   "EMP IDB_stations_me{16}_partNumbers{2}" : WString[40] = PLC "EMP IDB".stations.me[16].partNumbers[2], 1 s
   "EMP IDB_stations_me{16}_partNumbers{3}" : WString[40] = PLC "EMP IDB".stations.me[16].partNumbers[3], 1 s
   "EMP IDB_stations_me{16}_partNumbers{4}" : WString[40] = PLC "EMP IDB".stations.me[16].partNumbers[4], 1 s
   "EMP IDB_stations_me{16}_partNumbers{5}" : WString[40] = PLC "EMP IDB".stations.me[16].partNumbers[5], 1 s
   "EMP IDB_stations_me{16}_partNumbers{6}" : WString[40] = PLC "EMP IDB".stations.me[16].partNumbers[6], 1 s
   "EMP IDB_stations_me{16}_partNumbers{7}" : WString[40] = PLC "EMP IDB".stations.me[16].partNumbers[7], 1 s
   "EMP IDB_stations_me{17}_partNumbers{0}" : WString[40] = PLC "EMP IDB".stations.me[17].partNumbers[0], 1 s
   "EMP IDB_stations_me{17}_partNumbers{1}" : WString[40] = PLC "EMP IDB".stations.me[17].partNumbers[1], 1 s
   "EMP IDB_stations_me{17}_partNumbers{2}" : WString[40] = PLC "EMP IDB".stations.me[17].partNumbers[2], 1 s
   "EMP IDB_stations_me{17}_partNumbers{3}" : WString[40] = PLC "EMP IDB".stations.me[17].partNumbers[3], 1 s
   "EMP IDB_stations_me{17}_partNumbers{4}" : WString[40] = PLC "EMP IDB".stations.me[17].partNumbers[4], 1 s
   "EMP IDB_stations_me{17}_partNumbers{5}" : WString[40] = PLC "EMP IDB".stations.me[17].partNumbers[5], 1 s
   "EMP IDB_stations_me{17}_partNumbers{6}" : WString[40] = PLC "EMP IDB".stations.me[17].partNumbers[6], 1 s
   "EMP IDB_stations_me{17}_partNumbers{7}" : WString[40] = PLC "EMP IDB".stations.me[17].partNumbers[7], 1 s
   "EMP IDB_stations_me{18}_partNumbers{0}" : WString[40] = PLC "EMP IDB".stations.me[18].partNumbers[0], 1 s
   "EMP IDB_stations_me{18}_partNumbers{1}" : WString[40] = PLC "EMP IDB".stations.me[18].partNumbers[1], 1 s
   "EMP IDB_stations_me{18}_partNumbers{2}" : WString[40] = PLC "EMP IDB".stations.me[18].partNumbers[2], 1 s
   "EMP IDB_stations_me{18}_partNumbers{3}" : WString[40] = PLC "EMP IDB".stations.me[18].partNumbers[3], 1 s
   "EMP IDB_stations_me{18}_partNumbers{4}" : WString[40] = PLC "EMP IDB".stations.me[18].partNumbers[4], 1 s
   "EMP IDB_stations_me{18}_partNumbers{5}" : WString[40] = PLC "EMP IDB".stations.me[18].partNumbers[5], 1 s
   "EMP IDB_stations_me{18}_partNumbers{6}" : WString[40] = PLC "EMP IDB".stations.me[18].partNumbers[6], 1 s
   "EMP IDB_stations_me{18}_partNumbers{7}" : WString[40] = PLC "EMP IDB".stations.me[18].partNumbers[7], 1 s
   "EMP IDB_stations_me{19}_partNumbers{0}" : WString[40] = PLC "EMP IDB".stations.me[19].partNumbers[0], 1 s
   "EMP IDB_stations_me{19}_partNumbers{1}" : WString[40] = PLC "EMP IDB".stations.me[19].partNumbers[1], 1 s
   "EMP IDB_stations_me{19}_partNumbers{2}" : WString[40] = PLC "EMP IDB".stations.me[19].partNumbers[2], 1 s
   "EMP IDB_stations_me{19}_partNumbers{3}" : WString[40] = PLC "EMP IDB".stations.me[19].partNumbers[3], 1 s
   "EMP IDB_stations_me{19}_partNumbers{4}" : WString[40] = PLC "EMP IDB".stations.me[19].partNumbers[4], 1 s
   "EMP IDB_stations_me{19}_partNumbers{5}" : WString[40] = PLC "EMP IDB".stations.me[19].partNumbers[5], 1 s
   "EMP IDB_stations_me{19}_partNumbers{6}" : WString[40] = PLC "EMP IDB".stations.me[19].partNumbers[6], 1 s
   "EMP IDB_stations_me{19}_partNumbers{7}" : WString[40] = PLC "EMP IDB".stations.me[19].partNumbers[7], 1 s
   "EMP IDB_stations_me{20}_partNumbers{0}" : WString[40] = PLC "EMP IDB".stations.me[20].partNumbers[0], 1 s
   "EMP IDB_stations_me{20}_partNumbers{1}" : WString[40] = PLC "EMP IDB".stations.me[20].partNumbers[1], 1 s
   "EMP IDB_stations_me{20}_partNumbers{2}" : WString[40] = PLC "EMP IDB".stations.me[20].partNumbers[2], 1 s
   "EMP IDB_stations_me{20}_partNumbers{3}" : WString[40] = PLC "EMP IDB".stations.me[20].partNumbers[3], 1 s
   "EMP IDB_stations_me{20}_partNumbers{4}" : WString[40] = PLC "EMP IDB".stations.me[20].partNumbers[4], 1 s
   "EMP IDB_stations_me{20}_partNumbers{5}" : WString[40] = PLC "EMP IDB".stations.me[20].partNumbers[5], 1 s
   "EMP IDB_stations_me{20}_partNumbers{6}" : WString[40] = PLC "EMP IDB".stations.me[20].partNumbers[6], 1 s
   "EMP IDB_stations_me{20}_partNumbers{7}" : WString[40] = PLC "EMP IDB".stations.me[20].partNumbers[7], 1 s
   "EMP IDB_stations_me{21}_partNumbers{0}" : WString[40] = PLC "EMP IDB".stations.me[21].partNumbers[0], 1 s
   "EMP IDB_stations_me{21}_partNumbers{1}" : WString[40] = PLC "EMP IDB".stations.me[21].partNumbers[1], 1 s
   "EMP IDB_stations_me{21}_partNumbers{2}" : WString[40] = PLC "EMP IDB".stations.me[21].partNumbers[2], 1 s
   "EMP IDB_stations_me{21}_partNumbers{3}" : WString[40] = PLC "EMP IDB".stations.me[21].partNumbers[3], 1 s
   "EMP IDB_stations_me{21}_partNumbers{4}" : WString[40] = PLC "EMP IDB".stations.me[21].partNumbers[4], 1 s
   "EMP IDB_stations_me{21}_partNumbers{5}" : WString[40] = PLC "EMP IDB".stations.me[21].partNumbers[5], 1 s
   "EMP IDB_stations_me{21}_partNumbers{6}" : WString[40] = PLC "EMP IDB".stations.me[21].partNumbers[6], 1 s
   "EMP IDB_stations_me{21}_partNumbers{7}" : WString[40] = PLC "EMP IDB".stations.me[21].partNumbers[7], 1 s
   "EMP IDB_stations_me{22}_partNumbers{0}" : WString[40] = PLC "EMP IDB".stations.me[22].partNumbers[0], 1 s
   "EMP IDB_stations_me{22}_partNumbers{1}" : WString[40] = PLC "EMP IDB".stations.me[22].partNumbers[1], 1 s
   "EMP IDB_stations_me{22}_partNumbers{2}" : WString[40] = PLC "EMP IDB".stations.me[22].partNumbers[2], 1 s
   "EMP IDB_stations_me{22}_partNumbers{3}" : WString[40] = PLC "EMP IDB".stations.me[22].partNumbers[3], 1 s
   "EMP IDB_stations_me{22}_partNumbers{4}" : WString[40] = PLC "EMP IDB".stations.me[22].partNumbers[4], 1 s
   "EMP IDB_stations_me{22}_partNumbers{5}" : WString[40] = PLC "EMP IDB".stations.me[22].partNumbers[5], 1 s
   "EMP IDB_stations_me{22}_partNumbers{6}" : WString[40] = PLC "EMP IDB".stations.me[22].partNumbers[6], 1 s
   "EMP IDB_stations_me{22}_partNumbers{7}" : WString[40] = PLC "EMP IDB".stations.me[22].partNumbers[7], 1 s
   "EMP IDB_stations_me{23}_partNumbers{0}" : WString[40] = PLC "EMP IDB".stations.me[23].partNumbers[0], 1 s
   "EMP IDB_stations_me{23}_partNumbers{1}" : WString[40] = PLC "EMP IDB".stations.me[23].partNumbers[1], 1 s
   "EMP IDB_stations_me{23}_partNumbers{2}" : WString[40] = PLC "EMP IDB".stations.me[23].partNumbers[2], 1 s
   "EMP IDB_stations_me{23}_partNumbers{3}" : WString[40] = PLC "EMP IDB".stations.me[23].partNumbers[3], 1 s
   "EMP IDB_stations_me{23}_partNumbers{4}" : WString[40] = PLC "EMP IDB".stations.me[23].partNumbers[4], 1 s
   "EMP IDB_stations_me{23}_partNumbers{5}" : WString[40] = PLC "EMP IDB".stations.me[23].partNumbers[5], 1 s
   "EMP IDB_stations_me{23}_partNumbers{6}" : WString[40] = PLC "EMP IDB".stations.me[23].partNumbers[6], 1 s
   "EMP IDB_stations_me{23}_partNumbers{7}" : WString[40] = PLC "EMP IDB".stations.me[23].partNumbers[7], 1 s
   "EMP IDB_stations_me{3}_partNumbers{0}" : WString[40] = PLC "EMP IDB".stations.me[3].partNumbers[0], 1 s

text list "Station Selection Single": 0 'Select a Station to View'; 1 'Assignments'

recipe "VOLVO 16 01": Button 0 <- "EMP IDB_stations_me{0}_partNumbers{0}", Button 1 <- "EMP IDB_stations_me{0}_partNumbers{1}", Button 2 <- "EMP IDB_stations_me{0}_partNumbers{2}", Button 3 <- "EMP IDB_stations_me{0}_partNumbers{3}", Button 4 <- "EMP IDB_stations_me{0}_partNumbers{4}", Button 5 <- "EMP IDB_stations_me{0}_partNumbers{5}", Button 6 <- "EMP IDB_stations_me{0}_partNumbers{6}", Button 7 <- "EMP IDB_stations_me{0}_partNumbers{7}"

recipe "VOLVO 16 02": Button 0 <- "EMP IDB_stations_me{1}_partNumbers{0}", Button 1 <- "EMP IDB_stations_me{1}_partNumbers{1}", Button 2 <- "EMP IDB_stations_me{1}_partNumbers{2}", Button 3 <- "EMP IDB_stations_me{1}_partNumbers{3}", Button 4 <- "EMP IDB_stations_me{1}_partNumbers{4}", Button 5 <- "EMP IDB_stations_me{1}_partNumbers{5}", Button 6 <- "EMP IDB_stations_me{1}_partNumbers{6}", Button 7 <- "EMP IDB_stations_me{1}_partNumbers{7}"

recipe "VOLVO 16 03": Button 0 <- "EMP IDB_stations_me{2}_partNumbers{0}", Button 1 <- "EMP IDB_stations_me{2}_partNumbers{1}", Button 2 <- "EMP IDB_stations_me{2}_partNumbers{2}", Button 3 <- "EMP IDB_stations_me{2}_partNumbers{3}", Button 4 <- "EMP IDB_stations_me{2}_partNumbers{4}", Button 5 <- "EMP IDB_stations_me{2}_partNumbers{5}", Button 6 <- "EMP IDB_stations_me{2}_partNumbers{6}", Button 7 <- "EMP IDB_stations_me{2}_partNumbers{7}"

recipe "VOLVO 16 04": Button 0 <- "EMP IDB_stations_me{3}_partNumbers{0}", Button 1, Button 2, Button 3, Button 4, Button 5, Button 6, Button 7, Recipe_element_1

recipe "VOLVO 16 05": Button 0 <- "EMP IDB_stations_me{4}_partNumbers{0}", Button 1 <- "EMP IDB_stations_me{4}_partNumbers{1}", Button 2 <- "EMP IDB_stations_me{4}_partNumbers{2}", Button 3 <- "EMP IDB_stations_me{4}_partNumbers{3}", Button 4 <- "EMP IDB_stations_me{4}_partNumbers{4}", Button 5 <- "EMP IDB_stations_me{4}_partNumbers{5}", Button 6 <- "EMP IDB_stations_me{4}_partNumbers{6}", Button 7 <- "EMP IDB_stations_me{4}_partNumbers{7}"

recipe "VOLVO 16 06": Button 0 <- "EMP IDB_stations_me{5}_partNumbers{0}", Button 1 <- "EMP IDB_stations_me{5}_partNumbers{1}", Button 2 <- "EMP IDB_stations_me{5}_partNumbers{2}", Button 3 <- "EMP IDB_stations_me{5}_partNumbers{3}", Button 4 <- "EMP IDB_stations_me{5}_partNumbers{4}", Button 5 <- "EMP IDB_stations_me{5}_partNumbers{5}", Button 6 <- "EMP IDB_stations_me{5}_partNumbers{6}", Button 7 <- "EMP IDB_stations_me{5}_partNumbers{7}"

recipe "VOLVO 16 07": Button 0 <- "EMP IDB_stations_me{6}_partNumbers{0}", Button 1 <- "EMP IDB_stations_me{6}_partNumbers{1}", Button 2 <- "EMP IDB_stations_me{6}_partNumbers{2}", Button 3 <- "EMP IDB_stations_me{6}_partNumbers{3}", Button 4 <- "EMP IDB_stations_me{6}_partNumbers{4}", Button 5 <- "EMP IDB_stations_me{6}_partNumbers{5}", Button 6 <- "EMP IDB_stations_me{6}_partNumbers{6}", Button 7 <- "EMP IDB_stations_me{6}_partNumbers{7}"

recipe "VOLVO 16 08": Button 0 <- "EMP IDB_stations_me{7}_partNumbers{0}", Button 1 <- "EMP IDB_stations_me{7}_partNumbers{1}", Button 2 <- "EMP IDB_stations_me{7}_partNumbers{2}", Button 3 <- "EMP IDB_stations_me{7}_partNumbers{3}", Button 4 <- "EMP IDB_stations_me{7}_partNumbers{4}", Button 5 <- "EMP IDB_stations_me{7}_partNumbers{5}", Button 6 <- "EMP IDB_stations_me{7}_partNumbers{6}", Button 7 <- "EMP IDB_stations_me{7}_partNumbers{7}"

recipe "VOLVO 16 09": Button 0 <- "EMP IDB_stations_me{8}_partNumbers{0}", Button 1 <- "EMP IDB_stations_me{8}_partNumbers{1}", Button 2 <- "EMP IDB_stations_me{8}_partNumbers{2}", Button 3 <- "EMP IDB_stations_me{8}_partNumbers{3}", Button 4 <- "EMP IDB_stations_me{8}_partNumbers{4}", Button 5 <- "EMP IDB_stations_me{8}_partNumbers{5}", Button 6 <- "EMP IDB_stations_me{8}_partNumbers{6}", Button 7 <- "EMP IDB_stations_me{8}_partNumbers{7}"

recipe "VOLVO 16 10": Button 0 <- "EMP IDB_stations_me{9}_partNumbers{0}", Button 1 <- "EMP IDB_stations_me{9}_partNumbers{1}", Button 2 <- "EMP IDB_stations_me{9}_partNumbers{2}", Button 3 <- "EMP IDB_stations_me{9}_partNumbers{3}", Button 4 <- "EMP IDB_stations_me{9}_partNumbers{4}", Button 5 <- "EMP IDB_stations_me{9}_partNumbers{5}", Button 6 <- "EMP IDB_stations_me{9}_partNumbers{6}", Button 7 <- "EMP IDB_stations_me{9}_partNumbers{7}"

recipe "VOLVO 16 11": Button 0 <- "EMP IDB_stations_me{10}_partNumbers{0}", Button 1 <- "EMP IDB_stations_me{10}_partNumbers{1}", Button 2 <- "EMP IDB_stations_me{10}_partNumbers{2}", Button 3 <- "EMP IDB_stations_me{10}_partNumbers{3}", Button 4 <- "EMP IDB_stations_me{10}_partNumbers{4}", Button 5 <- "EMP IDB_stations_me{10}_partNumbers{5}", Button 6 <- "EMP IDB_stations_me{10}_partNumbers{6}", Button 7 <- "EMP IDB_stations_me{10}_partNumbers{7}"

recipe "CHM 01": Button 0 <- "EMP IDB_stations_me{11}_partNumbers{0}", Button 1 <- "EMP IDB_stations_me{11}_partNumbers{1}", Button 2 <- "EMP IDB_stations_me{11}_partNumbers{2}", Button 3 <- "EMP IDB_stations_me{11}_partNumbers{3}", Button 4 <- "EMP IDB_stations_me{11}_partNumbers{4}", Button 5 <- "EMP IDB_stations_me{11}_partNumbers{5}", Button 6 <- "EMP IDB_stations_me{11}_partNumbers{6}", Button 7 <- "EMP IDB_stations_me{11}_partNumbers{7}"

recipe "CHM 02": Button 0 <- "EMP IDB_stations_me{12}_partNumbers{0}", Button 1 <- "EMP IDB_stations_me{12}_partNumbers{1}", Button 2 <- "EMP IDB_stations_me{12}_partNumbers{2}", Button 3 <- "EMP IDB_stations_me{12}_partNumbers{3}", Button 4 <- "EMP IDB_stations_me{12}_partNumbers{4}", Button 5 <- "EMP IDB_stations_me{12}_partNumbers{5}", Button 6 <- "EMP IDB_stations_me{12}_partNumbers{6}", Button 7 <- "EMP IDB_stations_me{12}_partNumbers{7}"

recipe "CHM 03": Button 0 <- "EMP IDB_stations_me{13}_partNumbers{0}", Button 1 <- "EMP IDB_stations_me{13}_partNumbers{1}", Button 2 <- "EMP IDB_stations_me{13}_partNumbers{2}", Button 3 <- "EMP IDB_stations_me{13}_partNumbers{3}", Button 4 <- "EMP IDB_stations_me{13}_partNumbers{4}", Button 5 <- "EMP IDB_stations_me{13}_partNumbers{5}", Button 6 <- "EMP IDB_stations_me{13}_partNumbers{6}", Button 7 <- "EMP IDB_stations_me{13}_partNumbers{7}"

recipe "CHM 04": Button 0 <- "EMP IDB_stations_me{14}_partNumbers{0}", Button 1 <- "EMP IDB_stations_me{14}_partNumbers{1}", Button 2 <- "EMP IDB_stations_me{14}_partNumbers{2}", Button 3 <- "EMP IDB_stations_me{14}_partNumbers{3}", Button 4 <- "EMP IDB_stations_me{14}_partNumbers{4}", Button 5 <- "EMP IDB_stations_me{14}_partNumbers{5}", Button 6 <- "EMP IDB_stations_me{14}_partNumbers{6}", Button 7 <- "EMP IDB_stations_me{14}_partNumbers{7}"

recipe "CHM 05": Button 0 <- "EMP IDB_stations_me{15}_partNumbers{0}", Button 1 <- "EMP IDB_stations_me{15}_partNumbers{1}", Button 2 <- "EMP IDB_stations_me{15}_partNumbers{2}", Button 3 <- "EMP IDB_stations_me{15}_partNumbers{3}", Button 4 <- "EMP IDB_stations_me{15}_partNumbers{4}", Button 5 <- "EMP IDB_stations_me{15}_partNumbers{5}", Button 6 <- "EMP IDB_stations_me{15}_partNumbers{6}", Button 7 <- "EMP IDB_stations_me{15}_partNumbers{7}"

recipe "CDO 01": Button 0 <- "EMP IDB_stations_me{16}_partNumbers{0}", Button 1 <- "EMP IDB_stations_me{16}_partNumbers{1}", Button 2 <- "EMP IDB_stations_me{16}_partNumbers{2}", Button 3 <- "EMP IDB_stations_me{16}_partNumbers{3}", Button 4 <- "EMP IDB_stations_me{16}_partNumbers{4}", Button 5 <- "EMP IDB_stations_me{16}_partNumbers{5}", Button 6 <- "EMP IDB_stations_me{16}_partNumbers{6}", Button 7 <- "EMP IDB_stations_me{16}_partNumbers{7}"

recipe "CDO 02": Button 0 <- "EMP IDB_stations_me{17}_partNumbers{0}", Button 1 <- "EMP IDB_stations_me{17}_partNumbers{1}", Button 2 <- "EMP IDB_stations_me{17}_partNumbers{2}", Button 3 <- "EMP IDB_stations_me{17}_partNumbers{3}", Button 4 <- "EMP IDB_stations_me{17}_partNumbers{4}", Button 5 <- "EMP IDB_stations_me{17}_partNumbers{5}", Button 6 <- "EMP IDB_stations_me{17}_partNumbers{6}", Button 7 <- "EMP IDB_stations_me{17}_partNumbers{7}"

recipe "CDO 03": Button 0 <- "EMP IDB_stations_me{18}_partNumbers{0}", Button 1 <- "EMP IDB_stations_me{18}_partNumbers{1}", Button 2 <- "EMP IDB_stations_me{18}_partNumbers{2}", Button 3 <- "EMP IDB_stations_me{18}_partNumbers{3}", Button 4 <- "EMP IDB_stations_me{18}_partNumbers{4}", Button 5 <- "EMP IDB_stations_me{18}_partNumbers{5}", Button 6 <- "EMP IDB_stations_me{18}_partNumbers{6}", Button 7 <- "EMP IDB_stations_me{18}_partNumbers{7}"

recipe "BFL 01": Button 0 <- "EMP IDB_stations_me{19}_partNumbers{0}", Button 1 <- "EMP IDB_stations_me{19}_partNumbers{1}", Button 2 <- "EMP IDB_stations_me{19}_partNumbers{2}", Button 3 <- "EMP IDB_stations_me{19}_partNumbers{3}", Button 4 <- "EMP IDB_stations_me{19}_partNumbers{4}", Button 5 <- "EMP IDB_stations_me{19}_partNumbers{5}", Button 6 <- "EMP IDB_stations_me{19}_partNumbers{6}", Button 7 <- "EMP IDB_stations_me{19}_partNumbers{7}"

recipe "BFL 02": Button 0 <- "EMP IDB_stations_me{20}_partNumbers{0}", Button 1 <- "EMP IDB_stations_me{20}_partNumbers{1}", Button 2 <- "EMP IDB_stations_me{20}_partNumbers{2}", Button 3 <- "EMP IDB_stations_me{20}_partNumbers{3}", Button 4 <- "EMP IDB_stations_me{20}_partNumbers{4}", Button 5 <- "EMP IDB_stations_me{20}_partNumbers{5}", Button 6 <- "EMP IDB_stations_me{20}_partNumbers{6}", Button 7 <- "EMP IDB_stations_me{20}_partNumbers{7}"

recipe "BFL 03": Button 0 <- "EMP IDB_stations_me{21}_partNumbers{0}", Button 1 <- "EMP IDB_stations_me{21}_partNumbers{1}", Button 2 <- "EMP IDB_stations_me{21}_partNumbers{2}", Button 3 <- "EMP IDB_stations_me{21}_partNumbers{3}", Button 4 <- "EMP IDB_stations_me{21}_partNumbers{4}", Button 5 <- "EMP IDB_stations_me{21}_partNumbers{5}", Button 6 <- "EMP IDB_stations_me{21}_partNumbers{6}", Button 7 <- "EMP IDB_stations_me{21}_partNumbers{7}"

recipe "LGS 01": Button 0 <- "EMP IDB_stations_me{22}_partNumbers{0}", Button 1 <- "EMP IDB_stations_me{22}_partNumbers{1}", Button 2 <- "EMP IDB_stations_me{22}_partNumbers{2}", Button 3 <- "EMP IDB_stations_me{22}_partNumbers{3}", Button 4 <- "EMP IDB_stations_me{22}_partNumbers{4}", Button 5 <- "EMP IDB_stations_me{22}_partNumbers{5}", Button 6 <- "EMP IDB_stations_me{22}_partNumbers{6}", Button 7 <- "EMP IDB_stations_me{22}_partNumbers{7}"

recipe "LGS 02": Button 0 <- "EMP IDB_stations_me{23}_partNumbers{0}", Button 1 <- "EMP IDB_stations_me{23}_partNumbers{1}", Button 2 <- "EMP IDB_stations_me{23}_partNumbers{2}", Button 3 <- "EMP IDB_stations_me{23}_partNumbers{3}", Button 4 <- "EMP IDB_stations_me{23}_partNumbers{4}", Button 5 <- "EMP IDB_stations_me{23}_partNumbers{5}", Button 6 <- "EMP IDB_stations_me{23}_partNumbers{6}", Button 7 <- "EMP IDB_stations_me{23}_partNumbers{7}"

screen "1 PART CALL" 1366x768
   on GenerateScreen: SetTag("HMI_screenNumber", 1)
   Rectangle "Settings Tab Background" at 682,0 size 684x68
      Appearance <- "HMI_screenNumber"
   Rectangle "Part Call Tab Background" at 0,0 size 685x68
      Appearance <- "HMI_screenNumber"
   Rectangle "Settings Tab Border Hide" at 685,61 size 678x20
      Visibility <- "HMI_screenNumber"
   Rectangle "Part Call Tab Border Hide" at 3,61 size 679x20
      Visibility <- "HMI_screenNumber"
   Button "Settings Screen" at 683,0 size 683x68; TextOff 'SETTINGS'; Authorization "User administration"
      on Release: ActivateScreen("2 SETTINGS", 0)
   Button "Part Call Screen" at 0,0 size 683x68; TextOff 'PART CALL'
      on Release: ActivateScreen("1 PART CALL", 0)
   TextField "Header Line" at 32,112 size 216x53; Text 'LINE'
   TextField "Header Drop Zone" at 238,112 size 236x53; Text 'DROP ZONE'
   TextField "Header Part Number" at 474,112 size 648x53; Text 'PART NUMBER'
   TextField "Header Time" at 1112,112 size 222x53; Text 'TIME'
   ScreenModuleView "TableRow00" at 27,170 size 1312x52; ScreenModuleType ""
      Guid_{11997190-27688} <- "HMI_partCall_row{0}"
      on Guid_{11997190-83214}: ActivateScreen("3 BARCODE", 0)
   ScreenModuleView "TableRow01" at 27,222 size 1312x52; ScreenModuleType ""
      Guid_{11997190-27688} <- "HMI_partCall_row{1}"
      on Guid_{11997190-83214}: ActivateScreen("3 BARCODE", 0)
   ScreenModuleView "TableRow02" at 27,274 size 1312x52; ScreenModuleType ""
      Guid_{11997190-27688} <- "HMI_partCall_row{2}"
      on Guid_{11997190-83214}: ActivateScreen("3 BARCODE", 0)
   ScreenModuleView "TableRow03" at 27,326 size 1312x52; ScreenModuleType ""
      Guid_{11997190-27688} <- "HMI_partCall_row{3}"
      on Guid_{11997190-83214}: ActivateScreen("3 BARCODE", 0)
   ScreenModuleView "TableRow04" at 27,378 size 1312x52; ScreenModuleType ""
      Guid_{11997190-27688} <- "HMI_partCall_row{4}"
      on Guid_{11997190-83214}: ActivateScreen("3 BARCODE", 0)
   ScreenModuleView "TableRow05" at 27,430 size 1312x52; ScreenModuleType ""
      Guid_{11997190-27688} <- "HMI_partCall_row{5}"
      on Guid_{11997190-83214}: ActivateScreen("3 BARCODE", 0)
   ScreenModuleView "TableRow06" at 27,482 size 1312x52; ScreenModuleType ""
      Guid_{11997190-27688} <- "HMI_partCall_row{6}"
      on Guid_{11997190-83214}: ActivateScreen("3 BARCODE", 0)
   ScreenModuleView "TableRow07" at 27,534 size 1312x52; ScreenModuleType ""
      Guid_{11997190-27688} <- "HMI_partCall_row{7}"
      on Guid_{11997190-83214}: ActivateScreen("3 BARCODE", 0)
   ScreenModuleView "TableRow08" at 27,586 size 1312x52; ScreenModuleType ""
      Guid_{11997190-27688} <- "HMI_partCall_row{8}"
      on Guid_{11997190-83214}: ActivateScreen("3 BARCODE", 0)
   ScreenModuleView "TableRow09" at 27,638 size 1312x52; ScreenModuleType ""
      Guid_{11997190-27688} <- "HMI_partCall_row{9}"
      on Guid_{11997190-83214}: ActivateScreen("3 BARCODE", 0)
   ScreenModuleView "TableRow10" at 27,690 size 1312x52; ScreenModuleType ""
      Guid_{11997190-27688} <- "HMI_partCall_row{10}"
      on Guid_{11997190-83214}: ActivateScreen("3 BARCODE", 0)

screen "2 SETTINGS" 1366x768
   on GenerateScreen: SetTag("HMI_screenNumber", 2)
   Rectangle "Part Call Nave Panel" at 0,0 size 455x68
      Appearance <- "HMI_screenNumber"
   Rectangle "Settings Nav Panel" at 452,0 size 462x68
      Appearance <- "HMI_screenNumber"
   Rectangle "Network Health Nav Panel" at 911,0 size 455x68
      Appearance <- "HMI_screenNumber"
   Rectangle "Part Call Border Hide" at 3,60 size 449x20
      Visibility <- "HMI_screenNumber"
   Rectangle "Settings Border Hide" at 455,60 size 456x20
      Visibility <- "HMI_screenNumber"
   Rectangle "Network Health Border Hide" at 914,60 size 449x20
      Visibility <- "HMI_screenNumber"
   Button "Part Call Screen" at 0,0 size 455x68; TextOff 'PART CALL'
      on Release: ActivateScreen("1 PART CALL", 0)
   Button "Settings Screen" at 455,0 size 460x68; TextOff 'SETTINGS'
      on Release: ActivateScreen("2 SETTINGS", 0)
   Button "Network Health Screen" at 914,0 size 452x68; TextOff 'NW HEALTH'
      on Release: ActivateScreen("4 NETWORK HEALTH", 0)
   Rectangle "Station Assignment Table BG Full" at 793,120 size 533x630
      Visibility <- "HMI_settings_stations_selCount"
   TextField "Current Station Single" at 803,130 size 513x45; Text 'Text'
      Visibility <- "HMI_settings_stations_selCount"
   TextField "Hide Line and Drop Zone Multi" at 803,181 size 513x40; Text 'select single station for Line and Drop Zone'
      Visibility <- "HMI_settings_stations_selCount"
   GraphicView "KP8 Image" at 496,327 size 275x412; Picture "kp8 image"
   Rectangle "Station Assignment Table BG Mini" at 793,120 size 533x65
      Visibility <- "HMI_settings_stations_selCount"
   ScreenModuleView "PB: Set PN" at 50,130 size 414x45; Guid_{11997190-63616} 'Assign Part Number'; ScreenModuleType ""
      Guid_{11997190-63605} <- "HMI_settings_partNumber_assign"
   ScreenModuleView "PN IO Field" at 50,180 size 414x50; ScreenModuleType ""
      Guid_{11997190-63113} <- "HMI_settings_partNumber_ioField"
   ScreenModuleView "PB: Set Allotted" at 494,130 size 137x45; Guid_{11997190-63616} 'Allotted'; ScreenModuleType ""
      Guid_{11997190-63605} <- "HMI_settings_alotted_assign"
   ScreenModuleView "PB: Set Critical" at 636,130 size 137x45; Guid_{11997190-63616} 'Crititcal'; ScreenModuleType ""
      Guid_{11997190-63605} <- "HMI_settings_critical_assign"
   ScreenModuleView "Alotted Time IO Field" at 494,180 size 137x50; ScreenModuleType ""
      Guid_{11997190-63269} <- "HMI_settings_alotted_ioField"
   ScreenModuleView "Critical Time IO Field" at 636,180 size 137x50; ScreenModuleType ""
      Guid_{11997190-63269} <- "HMI_settings_critical_ioField"
   ScreenModuleView "PB: Select KP8 Buttons" at 493,270 size 284x45; Guid_{11997190-63616} 'Select Buttons'; ScreenModuleType ""
      Guid_{11997190-63605} <- "HMI_settings_kp8_selectButtons"
   ScreenModuleView "KP8 00: RESET" at 641,614 size 68x66; ScreenModuleType ""
      Guid_{11997190-57808} <- "HMI_settings_kp8_buttons{0}"
   ScreenModuleView "KP8 01" at 641,535 size 68x66; ScreenModuleType ""
      Guid_{11997190-57808} <- "HMI_settings_kp8_buttons{1}"
   ScreenModuleView "KP8 02" at 641,459 size 68x66; ScreenModuleType ""
      Guid_{11997190-57808} <- "HMI_settings_kp8_buttons{2}"
   ScreenModuleView "KP8 03" at 641,383 size 68x66; ScreenModuleType ""
      Guid_{11997190-57808} <- "HMI_settings_kp8_buttons{3}"
   ScreenModuleView "KP8 04: STOP RUNTIME" at 557,614 size 68x66; ScreenModuleType ""
      on Guid_{11997190-59171}: StopRuntime(0)
      Guid_{11997190-57808} <- "HMI_settings_kp8_buttons{4}"
   ScreenModuleView "KP8 05" at 557,535 size 68x66; ScreenModuleType ""
      Guid_{11997190-57808} <- "HMI_settings_kp8_buttons{5}"
   ScreenModuleView "KP8 06" at 557,459 size 68x66; ScreenModuleType ""
      Guid_{11997190-57808} <- "HMI_settings_kp8_buttons{6}"
   ScreenModuleView "KP8 07" at 557,383 size 68x66; ScreenModuleType ""
      Guid_{11997190-57808} <- "HMI_settings_kp8_buttons{7}"
   ScreenModuleView "PB: Previous Group" at 50,270 size 65x45; Guid_{11997190-63799} "Up"; ScreenModuleType ""
      Guid_{11997190-63779} <- "HMI_settings_stations_prevGroup"
   ScreenModuleView "PB: Select All Stations" at 120,270 size 274x45; Guid_{11997190-63616} 'Select Stations'; ScreenModuleType ""
      Guid_{11997190-63605} <- "HMI_settings_stations_selectAll"
   ScreenModuleView "PB: Next Group" at 399,270 size 65x45; Guid_{11997190-63799} "Down"; ScreenModuleType ""
      Guid_{11997190-63779} <- "HMI_settings_stations_nextGroup"
   ScreenModuleView "Station 00 Select" at 50,320 size 205x65; ScreenModuleType ""
      Guid_{11997190-57808} <- "HMI_settings_stations_selectBtns{0}"
   ScreenModuleView "Station 01 Select" at 260,320 size 205x65; ScreenModuleType ""
      Guid_{11997190-57808} <- "HMI_settings_stations_selectBtns{1}"
   ScreenModuleView "Station 02 Select" at 50,391 size 205x65; ScreenModuleType ""
      Guid_{11997190-57808} <- "HMI_settings_stations_selectBtns{2}"
   ScreenModuleView "Station 03 Select" at 260,391 size 205x65; ScreenModuleType ""
      Guid_{11997190-57808} <- "HMI_settings_stations_selectBtns{3}"
   ScreenModuleView "Station 04 Select" at 50,462 size 205x65; ScreenModuleType ""
      Guid_{11997190-57808} <- "HMI_settings_stations_selectBtns{4}"
   ScreenModuleView "Station 05 Select" at 260,462 size 205x65; ScreenModuleType ""
      Guid_{11997190-57808} <- "HMI_settings_stations_selectBtns{5}"
   ScreenModuleView "Station 06 Select" at 50,533 size 205x65; ScreenModuleType ""
      Guid_{11997190-57808} <- "HMI_settings_stations_selectBtns{6}"
   ScreenModuleView "Station 07 Select" at 260,533 size 205x65; ScreenModuleType ""
      Guid_{11997190-57808} <- "HMI_settings_stations_selectBtns{7}"
   ScreenModuleView "Station 08 Select" at 50,604 size 205x65; ScreenModuleType ""
      Guid_{11997190-57808} <- "HMI_settings_stations_selectBtns{8}"
   ScreenModuleView "Station 09 Select" at 260,604 size 205x65; ScreenModuleType ""
      Guid_{11997190-57808} <- "HMI_settings_stations_selectBtns{9}"
   ScreenModuleView "Station 10 Select" at 50,675 size 205x65; ScreenModuleType ""
      Guid_{11997190-57808} <- "HMI_settings_stations_selectBtns{10}"
   ScreenModuleView "Station 11 Select" at 260,675 size 205x65; ScreenModuleType ""
      Guid_{11997190-57808} <- "HMI_settings_stations_selectBtns{11}"
   ScreenModuleView "Line Label" at 803,181 size 267x40; ScreenModuleType ""
      Guid_{11997190-64598} <- "HMI_settings_viewingStation_lineData"
   ScreenModuleView "Drop Zone Label" at 1076,181 size 240x40; ScreenModuleType ""
      Guid_{11997190-64802} <- "HMI_settings_viewingStation_dzData"
   ScreenModuleView "PB: Previous Station" at 803,130 size 65x45; Guid_{11997190-63799} "Left"; ScreenModuleType ""
      Guid_{11997190-63779} <- "HMI_settings_viewingStation_previous"
   TextField "Current Station Multi" at 873,130 size 373x45; Text 'Assignments'
      Visibility <- "HMI_settings_stations_selCount"
   ScreenModuleView "PB: Next Station" at 1251,130 size 65x45; Guid_{11997190-63799} "Right"; ScreenModuleType ""
      Guid_{11997190-63779} <- "HMI_settings_viewingStation_next"
   TextField "Button Column Header" at 803,226 size 75x40; Text 'Btn'
      Visibility <- "HMI_settings_stations_selCount"
   TextField "Timer Column Header" at 872,226 size 128x40; Text 'Times'
      Visibility <- "HMI_settings_stations_selCount"
   TextField "Part Number Column Header" at 993,226 size 323x40; Text 'Part Number'
      Visibility <- "HMI_settings_stations_selCount"
   ScreenModuleView "Button 00 Details" at 803,271 size 513x74; ScreenModuleType ""
      Guid_{11997190-60358} <- "HMI_settings_viewingStation_btns{0}"
   ScreenModuleView "Button 01 Details" at 803,350 size 513x74; ScreenModuleType ""
      Guid_{11997190-60358} <- "HMI_settings_viewingStation_btns{1}"
   ScreenModuleView "Button 02 Details" at 803,429 size 513x74; ScreenModuleType ""
      Guid_{11997190-60358} <- "HMI_settings_viewingStation_btns{2}"
   ScreenModuleView "Button 03 Details" at 803,508 size 513x74; ScreenModuleType ""
      Guid_{11997190-60358} <- "HMI_settings_viewingStation_btns{3}"
   ScreenModuleView "Button 04 Details" at 803,587 size 513x74; ScreenModuleType ""
      Guid_{11997190-60358} <- "HMI_settings_viewingStation_btns{4}"
   ScreenModuleView "Button 05 Details" at 803,666 size 513x74; ScreenModuleType ""
      Guid_{11997190-60358} <- "HMI_settings_viewingStation_btns{5}"

SlideinScreen "GraphX_Slidein_Bottom" 1366x80
   ScreenModuleView "Top" at 0,0 size 227x80; Guid_{11997190-63799} "Top"; ScreenModuleType ""
      Guid_{11997190-63779} <- "HMI_tableNav_top"
   ScreenModuleView "Page Up" at 227,0 size 228x80; Guid_{11997190-63799} "pageUp"; ScreenModuleType ""
      Guid_{11997190-63779} <- "HMI_tableNav_pageUp"
   ScreenModuleView "Line Up" at 455,0 size 228x80; Guid_{11997190-63799} "Up"; ScreenModuleType ""
      Guid_{11997190-63779} <- "HMI_tableNav_lineUp"
   ScreenModuleView "Line Down" at 683,0 size 228x80; Guid_{11997190-63799} "Down"; ScreenModuleType ""
      Guid_{11997190-63779} <- "HMI_tableNav_lineDown"
   ScreenModuleView "Page Down" at 911,0 size 228x80; Guid_{11997190-63799} "PageDown"; ScreenModuleType ""
      Guid_{11997190-63779} <- "HMI_tableNav_pageDown"
   ScreenModuleView "Bottom" at 1138,0 size 228x80; Guid_{11997190-63799} "Bottom"; ScreenModuleType ""
      Guid_{11997190-63779} <- "HMI_tableNav_bottom"
   TextField "Text field_1" at 0,0 size 1366x80; Text 'NOT USED'
      Visibility <- "HMI_screenNumber"

SlideinScreen "GraphX_Slidein_Right" 449x768
   ScreenModuleView "Station Sim_1" at 5,5 size 106x232; ScreenModuleType ""
      Guid_{11997190-89108} <- "HMI_simStations_stations{0}"
   ScreenModuleView "Station Sim_2" at 116,5 size 106x232; ScreenModuleType ""
      Guid_{11997190-89108} <- "HMI_simStations_me{1}"
   ScreenModuleView "Station Sim_3" at 227,5 size 106x232; ScreenModuleType ""
      Guid_{11997190-89108} <- "HMI_simStations_me{2}"
   ScreenModuleView "Station Sim_4" at 338,5 size 106x232; ScreenModuleType ""
      Guid_{11997190-89108} <- "HMI_simStations_me{3}"
   ScreenModuleView "Station Sim_5" at 5,242 size 106x232; ScreenModuleType ""
      Guid_{11997190-89108} <- "HMI_simStations_me{4}"
   ScreenModuleView "Station Sim_6" at 5,479 size 106x232; ScreenModuleType ""
      Guid_{11997190-89108} <- "HMI_simStations_me{8}"
   ScreenModuleView "Station Sim_7" at 116,242 size 106x232; ScreenModuleType ""
      Guid_{11997190-89108} <- "HMI_simStations_me{5}"
   ScreenModuleView "Station Sim_8" at 227,242 size 106x232; ScreenModuleType ""
      Guid_{11997190-89108} <- "HMI_simStations_me{6}"
   ScreenModuleView "Station Sim_9" at 338,242 size 106x232; ScreenModuleType ""
      Guid_{11997190-89108} <- "HMI_simStations_me{7}"
   ScreenModuleView "Station Sim_10" at 116,479 size 106x232; ScreenModuleType ""
      Guid_{11997190-89108} <- "HMI_simStations_me{9}"
   ScreenModuleView "Station Sim_11" at 227,478 size 106x232; ScreenModuleType ""
      Guid_{11997190-89108} <- "HMI_simStations_me{10}"
   ScreenModuleView "Station Sim_12" at 338,477 size 106x232; ScreenModuleType ""
      Guid_{11997190-89108} <- "HMI_simStations_me{11}"
   ScreenModuleView "PB: Graphic/Text List_1" at 5,716 size 65x45; Guid_{11997190-63799} "Up"; ScreenModuleType ""
      Guid_{11997190-63779} <- "HMI_simStations_up"
   ScreenModuleView "PB: Graphic/Text List_2" at 379,716 size 65x45; Guid_{11997190-63799} "Down"; ScreenModuleType ""
      Guid_{11997190-63779} <- "HMI_simStations_down"

screen "3 BARCODE" 1366x768
   on GenerateScreen: SetTag("HMI_screenNumber", 3)
   Rectangle "Nav Panel 02" at 682,700 size 684x68
      Appearance <- "HMI_screenNumber"
   Rectangle "Nav Panel 01" at 0,700 size 685x68
      Appearance <- "HMI_screenNumber"
   Rectangle "Nav Panel 03 Top Border Hide" at 685,700 size 678x3
      Visibility <- "HMI_screenNumber"
   Rectangle "Nav Panel 01 Top Border Hide" at 3,700 size 679x3
      Visibility <- "HMI_screenNumber"
   Button "Settings Screen" at 683,700 size 683x68; TextOff 'SETTINGS'; Authorization "User administration"
      on Release: ActivateScreen("2 SETTINGS", 0)
   Button "Part Call Screen" at 0,700 size 683x68; TextOff 'PART CALL'
      on Release: ActivateScreen("1 PART CALL", 0)
   Button "btCancel" at 685,431 size 649x68; TextOff 'CANCEL'
      on Release: ActivateScreen("1 PART CALL", 0)
   Button "btPartOrdered" at 32,431 size 648x68; TextOff 'ORDERED'
      on Release: SetBit("ordered"); ActivateScreen("1 PART CALL", 0)
   TextField "tfBarcodeDisplay" at 32,220 size 1302x206; Text 'Text'
   TextField "tfPartNumberDisplay" at 32,160 size 1302x53; Text 'BARCODE FOR PART NUMBER'

screen "4 NETWORK HEALTH" 1366x768
   on GenerateScreen: SetTag("HMI_screenNumber", 4)
   ScreenModuleView "Volvo 16 Station 01 KP8" at 494,229 size 180x25; ScreenModuleType ""
      Guid_{11997190-57808} <- "HMI_networkHealth_pnioDevices{1}"
   ScreenModuleView "Volvo 16 Station 01 ET200SP" at 494,259 size 180x25; ScreenModuleType ""
      Guid_{11997190-57808} <- "HMI_networkHealth_pnioDevices{2}"
   ScreenModuleView "Volvo 16 Station 02 KP8" at 689,229 size 180x25; ScreenModuleType ""
      Guid_{11997190-57808} <- "HMI_networkHealth_pnioDevices{3}"
   ScreenModuleView "PB: Station Comm Status (Text Label)_4" at 689,259 size 180x25; ScreenModuleType ""
      Guid_{11997190-57808} <- "HMI_networkHealth_pnioDevices{4}"
   ScreenModuleView "PB: Station Comm Status (Text Label)_5" at 884,229 size 180x25; ScreenModuleType ""
      Guid_{11997190-57808} <- "HMI_networkHealth_pnioDevices{5}"
   ScreenModuleView "PB: Station Comm Status (Text Label)_6" at 884,259 size 180x25; ScreenModuleType ""
      Guid_{11997190-57808} <- "HMI_networkHealth_pnioDevices{6}"
   ScreenModuleView "PB: Station Comm Status (Text Label)_7" at 1079,229 size 180x25; ScreenModuleType ""
      Guid_{11997190-57808} <- "HMI_networkHealth_pnioDevices{7}"
   ScreenModuleView "PB: Station Comm Status (Text Label)_8" at 1079,259 size 180x25; ScreenModuleType ""
      Guid_{11997190-57808} <- "HMI_networkHealth_pnioDevices{8}"
   ScreenModuleView "PB: Station Comm Status (Text Label)_9" at 1079,154 size 180x25; ScreenModuleType ""
      Guid_{11997190-57808} <- "HMI_networkHealth_pnioDevices{9}"
   ScreenModuleView "PB: Station Comm Status (Text Label)_10" at 1079,184 size 180x25; ScreenModuleType ""
      Guid_{11997190-57808} <- "HMI_networkHealth_pnioDevices{10}"
   ScreenModuleView "PB: Station Comm Status (Text Label)_11" at 884,154 size 180x25; ScreenModuleType ""
      Guid_{11997190-57808} <- "HMI_networkHealth_pnioDevices{11}"
   ScreenModuleView "PB: Station Comm Status (Text Label)_12" at 884,184 size 180x25; ScreenModuleType ""
      Guid_{11997190-57808} <- "HMI_networkHealth_pnioDevices{12}"
   ScreenModuleView "PB: Station Comm Status (Text Label)_13" at 689,154 size 180x25; ScreenModuleType ""
      Guid_{11997190-57808} <- "HMI_networkHealth_pnioDevices{13}"
   ScreenModuleView "PB: Station Comm Status (Text Label)_14" at 689,184 size 180x25; ScreenModuleType ""
      Guid_{11997190-57808} <- "HMI_networkHealth_pnioDevices{14}"
   ScreenModuleView "PB: Station Comm Status (Text Label)_15" at 494,154 size 180x25; ScreenModuleType ""
      Guid_{11997190-57808} <- "HMI_networkHealth_pnioDevices{15}"
   ScreenModuleView "PB: Station Comm Status (Text Label)_16" at 494,184 size 180x25; ScreenModuleType ""
      Guid_{11997190-57808} <- "HMI_networkHealth_pnioDevices{16}"
   ScreenModuleView "PB: Station Comm Status (Text Label)_17" at 299,154 size 180x25; ScreenModuleType ""
      Guid_{11997190-57808} <- "HMI_networkHealth_pnioDevices{17}"
   ScreenModuleView "PB: Station Comm Status (Text Label)_18" at 299,184 size 180x25; ScreenModuleType ""
      Guid_{11997190-57808} <- "HMI_networkHealth_pnioDevices{18}"
   ScreenModuleView "PB: Station Comm Status (Text Label)_19" at 104,229 size 180x25; ScreenModuleType ""
      Guid_{11997190-57808} <- "HMI_networkHealth_pnioDevices{21}"
      on Guid_{11997190-101741}: SetTag("HMI_networkHealth_selectedDevice", 10)
   ScreenModuleView "PB: Station Comm Status (Text Label)_20" at 104,259 size 180x25; ScreenModuleType ""
      Guid_{11997190-57808} <- "HMI_networkHealth_pnioDevices{22}"
      on Guid_{11997190-101741}: SetTag("HMI_networkHealth_selectedDevice", 10)
   ScreenModuleView "PB: Station Comm Status (Text Label)_21" at 104,154 size 180x25; ScreenModuleType ""
      Guid_{11997190-57808} <- "HMI_networkHealth_pnioDevices{19}"
      on Guid_{11997190-101741}: function_efd93a16("KP8 Comm Status", 289, 40, -1, -1, 2); SetTag("HMI_networkHealth_selectedDevice", 10)
   ScreenModuleView "PB: Station Comm Status (Text Label)_22" at 104,184 size 180x25; ScreenModuleType ""
      Guid_{11997190-57808} <- "HMI_networkHealth_pnioDevices{20}"
      on Guid_{11997190-101741}: function_efd93a16("ET200SP Comm Status", 289, 40, -1, -1, 2); SetTag("HMI_networkHealth_selectedDevice", 10)
   ScreenModuleView "PB: Station Comm Status (Text Label)_23" at 105,323 size 180x25; ScreenModuleType ""
      Guid_{11997190-57808} <- "HMI_networkHealth_pnioDevices{31}"
   ScreenModuleView "PB: Station Comm Status (Text Label)_24" at 105,353 size 180x25; ScreenModuleType ""
      Guid_{11997190-57808} <- "HMI_networkHealth_pnioDevices{32}"
   ScreenModuleView "PB: Station Comm Status (Text Label)_25" at 299,323 size 180x25; ScreenModuleType ""
      Guid_{11997190-57808} <- "HMI_networkHealth_pnioDevices{29}"
   ScreenModuleView "PB: Station Comm Status (Text Label)_26" at 299,353 size 180x25; ScreenModuleType ""
      Guid_{11997190-57808} <- "HMI_networkHealth_pnioDevices{30}"
   ScreenModuleView "PB: Station Comm Status (Text Label)_27" at 105,396 size 180x25; ScreenModuleType ""
      Guid_{11997190-57808} <- "HMI_networkHealth_pnioDevices{23}"
   ScreenModuleView "PB: Station Comm Status (Text Label)_28" at 105,427 size 180x25; ScreenModuleType ""
      Guid_{11997190-57808} <- "HMI_networkHealth_pnioDevices{24}"
   ScreenModuleView "PB: Station Comm Status (Text Label)_29" at 299,396 size 180x25; ScreenModuleType ""
      Guid_{11997190-57808} <- "HMI_networkHealth_pnioDevices{27}"
   ScreenModuleView "PB: Station Comm Status (Text Label)_30" at 299,427 size 180x25; ScreenModuleType ""
      Guid_{11997190-57808} <- "HMI_networkHealth_pnioDevices{28}"
   ScreenModuleView "PB: Station Comm Status (Text Label)_31" at 105,468 size 180x25; ScreenModuleType ""
      Guid_{11997190-57808} <- "HMI_networkHealth_pnioDevices{25}"
   ScreenModuleView "PB: Station Comm Status (Text Label)_32" at 105,497 size 180x25; ScreenModuleType ""
      Guid_{11997190-57808} <- "HMI_networkHealth_pnioDevices{26}"
   ScreenModuleView "PB: Station Comm Status (Text Label)_33" at 105,558 size 180x25; ScreenModuleType ""
      Guid_{11997190-57808} <- "HMI_networkHealth_pnioDevices{33}"
   ScreenModuleView "PB: Station Comm Status (Text Label)_34" at 105,587 size 180x25; ScreenModuleType ""
      Guid_{11997190-57808} <- "HMI_networkHealth_pnioDevices{34}"
   ScreenModuleView "PB: Station Comm Status (Text Label)_35" at 105,623 size 180x25; ScreenModuleType ""
      Guid_{11997190-57808} <- "HMI_networkHealth_pnioDevices{37}"
   ScreenModuleView "PB: Station Comm Status (Text Label)_36" at 105,651 size 180x25; ScreenModuleType ""
      Guid_{11997190-57808} <- "HMI_networkHealth_pnioDevices{38}"
   ScreenModuleView "PB: Station Comm Status (Text Label)_37" at 299,558 size 180x25; ScreenModuleType ""
      Guid_{11997190-57808} <- "HMI_networkHealth_pnioDevices{35}"
   ScreenModuleView "PB: Station Comm Status (Text Label)_38" at 299,587 size 180x25; ScreenModuleType ""
      Guid_{11997190-57808} <- "HMI_networkHealth_pnioDevices{36}"
   ScreenModuleView "PB: Station Comm Status (Text Label)_39" at 103,691 size 180x25; ScreenModuleType ""
      Guid_{11997190-57808} <- "HMI_networkHealth_pnioDevices{43}"
   ScreenModuleView "PB: Station Comm Status (Text Label)_40" at 103,720 size 180x25; ScreenModuleType ""
      Guid_{11997190-57808} <- "HMI_networkHealth_pnioDevices{44}"
   ScreenModuleView "PB: Station Comm Status (Text Label)_41" at 298,627 size 180x25; ScreenModuleType ""
      Guid_{11997190-57808} <- "HMI_networkHealth_pnioDevices{39}"
   ScreenModuleView "PB: Station Comm Status (Text Label)_42" at 298,655 size 180x25; ScreenModuleType ""
      Guid_{11997190-57808} <- "HMI_networkHealth_pnioDevices{40}"
   ScreenModuleView "PB: Station Comm Status (Text Label)_43" at 297,691 size 180x25; ScreenModuleType ""
      Guid_{11997190-57808} <- "HMI_networkHealth_pnioDevices{41}"
   ScreenModuleView "PB: Station Comm Status (Text Label)_44" at 297,720 size 180x25; ScreenModuleType ""
      Guid_{11997190-57808} <- "HMI_networkHealth_pnioDevices{42}"
   ScreenModuleView "PB: Station Comm Status (Text Label)_45" at 495,324 size 180x25; ScreenModuleType ""
      Guid_{11997190-57808} <- "HMI_networkHealth_pnioDevices{45}"
   ScreenModuleView "PB: Station Comm Status (Text Label)_46" at 495,354 size 180x25; ScreenModuleType ""
      Guid_{11997190-57808} <- "HMI_networkHealth_pnioDevices{46}"
   ScreenModuleView "PB: Station Comm Status (Text Label)_47" at 689,397 size 180x25; ScreenModuleType ""
      Guid_{11997190-57808} <- "HMI_networkHealth_pnioDevices{47}"
   ScreenModuleView "PB: Station Comm Status (Text Label)_48" at 689,428 size 180x25; ScreenModuleType ""
      Guid_{11997190-57808} <- "HMI_networkHealth_pnioDevices{48}"
   Rectangle "Part Call Nave Panel" at 0,0 size 455x68
      Appearance <- "HMI_screenNumber"
   Rectangle "Settings Nav Panel" at 452,0 size 462x68
      Appearance <- "HMI_screenNumber"
   Rectangle "Network Health Nav Panel" at 911,0 size 455x68
      Appearance <- "HMI_screenNumber"
   Rectangle "Part Call Border Hide" at 3,60 size 449x20
      Visibility <- "HMI_screenNumber"
   Rectangle "Settings Border Hide" at 455,60 size 456x20
      Visibility <- "HMI_screenNumber"
   Rectangle "Network Health Border Hide" at 914,60 size 449x20
      Visibility <- "HMI_screenNumber"
   Button "Part Call Screen" at 0,0 size 455x68; TextOff 'PART CALL'
      on Release: ActivateScreen("1 PART CALL", 0)
   Button "Settings Screen" at 455,0 size 460x68; TextOff 'SETTINGS'
      on Release: ActivateScreen("2 SETTINGS", 0)
   Button "Network Health Screen" at 914,0 size 452x68; TextOff 'NW HEALTH'
      on Release: ActivateScreen("4 NETWORK HEALTH", 0)

PopupScreen "KP8 Comm Status" 438x720
   ScreenModuleView "Station: KP8_1" at 5,5 size 428x710; ScreenModuleType ""
      Guid_{11997190-107144} <- "HMI_networkHealth_kp8PopUp"
      on Guid_{11997190-107182}: function_efd93a16("KP8 Comm Status", 0, 0, -1, -1, 1)

PopupScreen "ET200SP Comm Status" 613x720
   ScreenModuleView "Station: ET200SP_1" at 5,5 size 603x710; ScreenModuleType ""
      Guid_{11997190-102952} <- "HMI_networkHealth_et200spPopUp"
      on Guid_{11997190-102950}: function_efd93a16("ET200SP Comm Status", 0, 0, -1, -1, 1)
*)

(* ===== HMI "HMI_RT_2" =====
connection "HMI_Connection_3": ETHERNET, S7_1500_OMS

HMI tags "Default tag table"
   "Clock_0.5Hz" : Bool = PLC "Clock_0.5Hz" AT %M0.7, 100 ms
   "LED Sign_request_row{0}" : Table Row = PLC "LED Sign".request.row[0], 100 ms
   "LED Sign_request_row{1}" : Table Row = PLC "LED Sign".request.row[1], 100 ms
   "LED Sign_request_row{2}" : Table Row = PLC "LED Sign".request.row[2], 100 ms
   "LED Sign_request_row{3}" : Table Row = PLC "LED Sign".request.row[3], 100 ms
   "LED Sign_request_row{4}" : Table Row = PLC "LED Sign".request.row[4], 100 ms
   "LED Sign_request_row{5}" : Table Row = PLC "LED Sign".request.row[5], 100 ms
   "LED Sign_request_row{6}" : Table Row = PLC "LED Sign".request.row[6], 100 ms
   "LED Sign_request_row{7}" : Table Row = PLC "LED Sign".request.row[7], 100 ms
   "LED Sign_request_row{8}" : Table Row = PLC "LED Sign".request.row[8], 100 ms
   "LED Sign_request_row{9}" : Table Row = PLC "LED Sign".request.row[9], 100 ms
   "LED Sign_request_row{10}" : Table Row = PLC "LED Sign".request.row[10], 100 ms
   "LED Sign_request_row{11}" : Table Row = PLC "LED Sign".request.row[11], 100 ms

screen "1 PART CALL" 1024x768
   Rectangle "Connection Status" at 1,196 size 894x1
      Appearance <- "Clock_0.5Hz"
   ScreenModuleView "R0C0" at 6,9 size 440x28; ScreenModuleType ""
      Guid_{11997190-27688} <- "LED Sign_request_row{0}"
   ScreenModuleView "R1C0" at 6,39 size 440x28; ScreenModuleType ""
      Guid_{11997190-27688} <- "LED Sign_request_row{1}"
   ScreenModuleView "R2C0" at 6,69 size 440x28; ScreenModuleType ""
      Guid_{11997190-27688} <- "LED Sign_request_row{2}"
   ScreenModuleView "R3C0" at 6,99 size 440x28; ScreenModuleType ""
      Guid_{11997190-27688} <- "LED Sign_request_row{3}"
   ScreenModuleView "R4C0" at 6,128 size 440x28; ScreenModuleType ""
      Guid_{11997190-27688} <- "LED Sign_request_row{4}"
   ScreenModuleView "R5C0" at 6,158 size 440x28; ScreenModuleType ""
      Guid_{11997190-27688} <- "LED Sign_request_row{5}"
   ScreenModuleView "R0C1" at 455,9 size 438x28; ScreenModuleType ""
      Guid_{11997190-27688} <- "LED Sign_request_row{6}"
   ScreenModuleView "R1C1" at 455,39 size 438x28; ScreenModuleType ""
      Guid_{11997190-27688} <- "LED Sign_request_row{7}"
   ScreenModuleView "R2C1" at 454,69 size 440x28; ScreenModuleType ""
      Guid_{11997190-27688} <- "LED Sign_request_row{8}"
   ScreenModuleView "R3C1" at 454,99 size 440x28; ScreenModuleType ""
      Guid_{11997190-27688} <- "LED Sign_request_row{9}"
   ScreenModuleView "R4C1" at 454,128 size 440x28; ScreenModuleType ""
      Guid_{11997190-27688} <- "LED Sign_request_row{10}"
   ScreenModuleView "R5C1" at 454,158 size 440x28; ScreenModuleType ""
      Guid_{11997190-27688} <- "LED Sign_request_row{11}"
*)

(* ===== HMI "HMI_RT_1" =====
system functions are stored by id; their names below are inferred from use

ScreenModuleEditorView "Table Row" 1312x52
   TextField "tfLine" at 5,1 size 216x48; Text 'Text'
      Visibility <- "interface.tfLine.visibility"
      Appearance <- "interface.tfLine.animator"
   TextField "tfTime" at 1085,1 size 222x48; Text 'Text'
      Appearance <- "interface.tfTime.animator"
      Visibility <- "interface.tfTime.visibility"
   TextField "tfDropZone" at 211,1 size 236x48; Text 'Text'
      Appearance <- "interface.tfDropZone.animator"
      Visibility <- "interface.tfDropZone.visibility"
   TextField "tfPartNumber" at 445,1 size 650x48; Text 'Text'
      Appearance <- "interface.tfPartNumber.animator"
      Visibility <- "interface.tfPartNumber.visibility"
   Button "pbSelect" at 0,0 size 1312x52; TextOff 'Text'
      Visibility <- "interface.pbSelection.visibility"
      on Press: SetBit("interface.pbSelection.request")
      on Release: ResetBit("interface.pbSelection.request")
   Rectangle "rtBackground" at 0,0 size 1312x52
      Visibility <- "interface.rtBackground.visibility"
*)

(* ===== HMI "HMI_RT_1" =====
system functions are stored by id; their names below are inferred from use

ScreenModuleEditorView "Table Row" 1312x52
   TextField "tfLine" at 5,1 size 216x48; Text 'Text'
      Visibility <- "interface.tfLine.visibility"
      Appearance <- "interface.tfLine.animator"
   TextField "tfTime" at 1085,1 size 222x48; Text 'Text'
      Visibility <- "interface.tfTime.visibility"
      Appearance <- "interface.tfTime.animator"
   TextField "tfDropZone" at 211,1 size 236x48; Text 'Text'
      Visibility <- "interface.tfDropZone.visibility"
      Appearance <- "interface.tfDropZone.animator"
   TextField "tfPartNumber" at 445,1 size 650x48; Text 'Text'
      Visibility <- "interface.tfPartNumber.visibility"
      Appearance <- "interface.tfPartNumber.animator"
   Button "pbSelect" at 0,0 size 1312x52; TextOff 'Text'
      on Release: ResetBit("interface.pbSelection.request")
      on Press: SetBit("interface.pbSelection.request")
      Visibility <- "interface.pbSelection.visibility"
   Rectangle "rtBackground" at 0,0 size 1312x52
      Visibility <- "interface.rtBackground.visibility"
*)

(* ===== HMI "HMI_RT_1" =====
system functions are stored by id; their names below are inferred from use

ScreenModuleEditorView "Table Row" 1312x52
   TextField "tfLine" at 5,1 size 216x48; Text 'Text'
      Visibility <- "interface.tfLine.visibility"
      Appearance <- "interface.tfLine.animator"
   TextField "tfTime" at 1085,1 size 222x48; Text 'Text'
      Visibility <- "interface.tfTime.visibility"
      Appearance <- "interface.tfTime.animator"
   TextField "tfDropZone" at 211,1 size 236x48; Text 'Text'
      Visibility <- "interface.tfDropZone.visibility"
      Appearance <- "interface.tfDropZone.animator"
   TextField "tfPartNumber" at 445,1 size 650x48; Text 'Text'
      Visibility <- "interface.tfPartNumber.visibility"
      Appearance <- "interface.tfPartNumber.animator"
   Button "pbSelect" at 0,0 size 1312x52; TextOff 'Text'
      on Release: ResetBit("interface.pbSelection.request")
      on Press: SetBit("interface.pbSelection.request")
      Visibility <- "interface.pbSelection.visibility"
   Rectangle "rtBackground" at 0,0 size 1312x52
      Visibility <- "interface.rtBackground.visibility"
*)

(* ===== HMI "HMI_RT_1" =====
system functions are stored by id; their names below are inferred from use

